
ScreenModuleEditorView "Station: ET200SP" 593x700
   GraphicView "ET200SP Stencil" at 0,50 size 593x649; Picture "ET 200SP Stencil"
   Rectangle "Interface Module Color" at 0,50 size 269x650
      Appearance <- "Interface.IM.bg"
   Rectangle "DQ 01 Module Color" at 268,50 size 95x344
      Appearance <- "Interface.DQ01.bg"
   Rectangle "DQ 01 Terminal Color" at 268,390 size 96x271
      Appearance <- "Interface.DQ01.bgTem"
   Rectangle "DQ 02 Module Color" at 363,50 size 96x344
      Appearance <- "Interface.DQ02.bg"
   Rectangle "DQ 02 Terminal Color" at 364,390 size 95x271
      Appearance <- "Interface.DQ02.bgTem"
   Rectangle "DQ 03 Module Color" at 458,50 size 95x344
      Appearance <- "Interface.DQ03.bg"
   Rectangle "DQ 03 Terminal Color" at 458,390 size 95x271
      Appearance <- "Interface.DQ03.bgTem"
   Rectangle "Server Module Color" at 552,50 size 40x343
      Appearance <- "Interface.serverModule.bg"
   Rectangle "IM Run LED" at 165,102 size 9x8
      Appearance <- "Interface.IM.run"
   Rectangle "IM Error LED" at 178,102 size 9x8
      Appearance <- "Interface.IM.error"
   Rectangle "IM Maintenance LED" at 193,102 size 9x8
      Appearance <- "Interface.IM.maint"
   Rectangle "IM Link 1 LED" at 146,295 size 9x8
      Appearance <- "Interface.IM.lnk01"
   Rectangle "IM Link 2 LED" at 146,313 size 9x8
      Appearance <- "Interface.IM.lnk02"
   Rectangle "IM Power LED" at 164,379 size 9x8
      Appearance <- "Interface.IM.pwr"
   Rectangle "DQ 01 Diag LED" at 274,102 size 9x8
      Appearance <- "Interface.DQ01.diag"
   Rectangle "DQ 01 Output LED x.0" at 274,295 size 9x8
      Appearance <- "Interface.DQ01.x0"
   Rectangle "DQ 01 Output LED x.1" at 305,295 size 9x8
      Appearance <- "Interface.DQ01.x1"
   Rectangle "DQ 01 Output LED x.2" at 274,306 size 9x8
      Appearance <- "Interface.DQ01.x2"
   Rectangle "DQ 01 Output LED x.3" at 305,306 size 9x8
      Appearance <- "Interface.DQ01.x3"
   Rectangle "DQ 01 Output LED x.4" at 274,317 size 9x8
      Appearance <- "Interface.DQ01.x4"
   Rectangle "DQ 01 Output LED x.5" at 305,317 size 9x8
      Appearance <- "Interface.DQ01.x5"
   Rectangle "DQ 01 Output LED x.6" at 274,328 size 9x8
      Appearance <- "Interface.DQ01.x6"
   Rectangle "DQ 01 Output LED x.7" at 305,328 size 9x8
      Appearance <- "Interface.DQ01.x7"
   Rectangle "DQ 01 Power LED" at 275,379 size 9x8
      Appearance <- "Interface.DQ01.pwr"
   Rectangle "DQ 02 Diag LED" at 369,102 size 9x8
      Appearance <- "Interface.DQ02.diag"
   Rectangle "DQ 02 Output LED x.0" at 369,295 size 9x8
      Appearance <- "Interface.DQ02.x0"
   Rectangle "DQ 02 Output LED x.1" at 400,295 size 9x8
      Appearance <- "Interface.DQ02.x1"
   Rectangle "DQ 02 Output LED x.2" at 369,306 size 9x8
      Appearance <- "Interface.DQ02.x2"
   Rectangle "DQ 02 Output LED x.3" at 400,306 size 9x8
      Appearance <- "Interface.DQ02.x3"
   Rectangle "DQ 02 Output LED x.4" at 369,317 size 9x8
      Appearance <- "Interface.DQ02.x4"
   Rectangle "DQ 02 Output LED x.5" at 400,317 size 9x8
      Appearance <- "Interface.DQ02.x5"
   Rectangle "DQ 02 Output LED x.6" at 369,328 size 9x8
      Appearance <- "Interface.DQ02.x6"
   Rectangle "DQ 02 Output LED x.7" at 400,328 size 9x8
      Appearance <- "Interface.DQ02.x7"
   Rectangle "DQ 02 Power LED" at 368,379 size 9x8
      Appearance <- "Interface.DQ02.pwr"
   Rectangle "DQ 03 Diag LED" at 464,102 size 9x8
      Appearance <- "Interface.DQ03.diag"
   Rectangle "DQ 03 Output LED x.0" at 464,295 size 9x8
      Appearance <- "Interface.DQ03.x0"
   Rectangle "DQ 03 Output LED x.1" at 495,295 size 9x8
      Appearance <- "Interface.DQ03.x1"
   Rectangle "DQ 03 Output LED x.2" at 464,306 size 9x8
      Appearance <- "Interface.DQ03.x2"
   Rectangle "DQ 03 Output LED x.3" at 495,306 size 9x8
      Appearance <- "Interface.DQ03.x3"
   Rectangle "DQ 03 Output LED x.4" at 464,317 size 9x8
      Appearance <- "Interface.DQ03.x4"
   Rectangle "DQ 03 Output LED x.5" at 495,317 size 9x8
      Appearance <- "Interface.DQ03.x5"
   Rectangle "DQ 03 Output LED x.6" at 464,328 size 9x8
      Appearance <- "Interface.DQ03.x6"
   Rectangle "DQ 03 Output LED x.7" at 495,328 size 9x8
      Appearance <- "Interface.DQ03.x7"
   Rectangle "DQ 03 Power LED" at 463,379 size 9x8
      Appearance <- "Interface.DQ03.pwr"
   Button "Dismiss PB" at 0,0 size 593x700; TextOff 'Text'
   TextField "PN Name" at 0,0 size 593x50; Text 'Text'
      Appearance <- "Interface.profinetName.animate"
*)

(* ===== HMI "HMI_RT_1" =====

ScreenModuleEditorView "Station: ET200SP" 603x710
   Rectangle "Interface Module Color" at 5,55 size 269x650
      Appearance <- "Interface.IM.bg"
   Rectangle "DQ 01 Module Color" at 273,55 size 95x344
      Appearance <- "Interface.DQ01.bg"
   Rectangle "DQ 01 Terminal Color" at 273,395 size 96x271
      Appearance <- "Interface.DQ01.bgTem"
   Rectangle "DQ 02 Module Color" at 368,55 size 96x344
      Appearance <- "Interface.DQ02.bg"
   Rectangle "DQ 02 Terminal Color" at 369,395 size 95x271
      Appearance <- "Interface.DQ02.bgTem"
   Rectangle "DQ 03 Module Color" at 463,55 size 95x344
      Appearance <- "Interface.DQ03.bg"
   Rectangle "DQ 03 Terminal Color" at 463,395 size 95x271
      Appearance <- "Interface.DQ03.bgTem"
   Rectangle "Server Module Color" at 557,55 size 40x343
      Appearance <- "Interface.serverModule.bg"
   Rectangle "IM Run LED" at 170,107 size 9x8
      Appearance <- "Interface.IM.run"
   Rectangle "IM Error LED" at 183,107 size 9x8
      Appearance <- "Interface.IM.error"
   Rectangle "IM Maintenance LED" at 198,107 size 9x8
      Appearance <- "Interface.IM.maint"
   Rectangle "IM Link 1 LED" at 151,300 size 9x8
      Appearance <- "Interface.IM.lnk01"
   Rectangle "IM Link 2 LED" at 151,318 size 9x8
      Appearance <- "Interface.IM.lnk02"
   Rectangle "IM Power LED" at 169,384 size 9x8
      Appearance <- "Interface.IM.pwr"
   Rectangle "DQ 01 Diag LED" at 279,107 size 9x8
      Appearance <- "Interface.DQ01.diag"
   Rectangle "DQ 01 Output LED x.0" at 279,300 size 9x8
      Appearance <- "Interface.DQ01.x0"
   Rectangle "DQ 01 Output LED x.1" at 310,300 size 9x8
      Appearance <- "Interface.DQ01.x1"
   Rectangle "DQ 01 Output LED x.2" at 279,311 size 9x8
      Appearance <- "Interface.DQ01.x2"
   Rectangle "DQ 01 Output LED x.3" at 310,311 size 9x8
      Appearance <- "Interface.DQ01.x3"
   Rectangle "DQ 01 Output LED x.4" at 279,322 size 9x8
      Appearance <- "Interface.DQ01.x4"
   Rectangle "DQ 01 Output LED x.5" at 310,322 size 9x8
      Appearance <- "Interface.DQ01.x5"
   Rectangle "DQ 01 Output LED x.6" at 279,333 size 9x8
      Appearance <- "Interface.DQ01.x6"
   Rectangle "DQ 01 Output LED x.7" at 310,333 size 9x8
      Appearance <- "Interface.DQ01.x7"
   Rectangle "DQ 01 Power LED" at 280,384 size 9x8
      Appearance <- "Interface.DQ01.pwr"
   Rectangle "DQ 02 Diag LED" at 374,107 size 9x8
      Appearance <- "Interface.DQ02.diag"
   Rectangle "DQ 02 Output LED x.0" at 374,300 size 9x8
      Appearance <- "Interface.DQ02.x0"
   Rectangle "DQ 02 Output LED x.1" at 405,300 size 9x8
      Appearance <- "Interface.DQ02.x1"
   Rectangle "DQ 02 Output LED x.2" at 374,311 size 9x8
      Appearance <- "Interface.DQ02.x2"
   Rectangle "DQ 02 Output LED x.3" at 405,311 size 9x8
      Appearance <- "Interface.DQ02.x3"
   Rectangle "DQ 02 Output LED x.4" at 374,322 size 9x8
      Appearance <- "Interface.DQ02.x4"
   Rectangle "DQ 02 Output LED x.5" at 405,322 size 9x8
      Appearance <- "Interface.DQ02.x5"
   Rectangle "DQ 02 Output LED x.6" at 374,333 size 9x8
      Appearance <- "Interface.DQ02.x6"
   Rectangle "DQ 02 Output LED x.7" at 405,333 size 9x8
      Appearance <- "Interface.DQ02.x7"
   Rectangle "DQ 02 Power LED" at 373,384 size 9x8
      Appearance <- "Interface.DQ02.pwr"
   Rectangle "DQ 03 Diag LED" at 469,107 size 9x8
      Appearance <- "Interface.DQ03.diag"
   Rectangle "DQ 03 Output LED x.0" at 469,300 size 9x8
      Appearance <- "Interface.DQ03.x0"
   Rectangle "DQ 03 Output LED x.1" at 500,300 size 9x8
      Appearance <- "Interface.DQ03.x1"
   Rectangle "DQ 03 Output LED x.2" at 469,311 size 9x8
      Appearance <- "Interface.DQ03.x2"
   Rectangle "DQ 03 Output LED x.3" at 500,311 size 9x8
      Appearance <- "Interface.DQ03.x3"
   Rectangle "DQ 03 Output LED x.4" at 469,322 size 9x8
      Appearance <- "Interface.DQ03.x4"
   Rectangle "DQ 03 Output LED x.5" at 500,322 size 9x8
      Appearance <- "Interface.DQ03.x5"
   Rectangle "DQ 03 Output LED x.6" at 469,333 size 9x8
      Appearance <- "Interface.DQ03.x6"
   Rectangle "DQ 03 Output LED x.7" at 500,333 size 9x8
      Appearance <- "Interface.DQ03.x7"
   Rectangle "DQ 03 Power LED" at 468,384 size 9x8
      Appearance <- "Interface.DQ03.pwr"
   GraphicView "ET200SP Stencil" at 5,55 size 593x649; Picture "ET 200SP Stencil"
   Button "Dismiss PB" at 5,5 size 593x700; TextOff 'Text'
   TextField "PN Name" at 5,5 size 593x50; Text 'Text'
      Appearance <- "Interface.profinetName.animate"
*)

(* ===== HMI "HMI_RT_1" =====

ScreenModuleEditorView "Station: KP8" 428x710
   GraphicView "KP8 Stencil" at 5,55 size 418x650; Picture "KP8 Rear View Stencil"
      Appearance <- "Interface.stencilBackground"
   TextField "PN Name Label" at 5,5 size 418x50; Text 'Text'
      Appearance <- "Interface.profinetName.animate"
   Rectangle "X1P1 Transmit" at 195,536 size 12x16
      Appearance <- "Interface.X1P1.transmit"
   Rectangle "X1P1 Receive" at 195,576 size 12x16
      Appearance <- "Interface.X1P1.receive"
   Rectangle "X1P2 Transmit" at 286,535 size 12x16
      Appearance <- "Interface.X1P2.transmit"
   Rectangle "X1P2 Receive" at 286,575 size 12x16
      Appearance <- "Interface.X1P2.receive"
   Rectangle "KP8 Background" at 5,55 size 418x650
      Appearance <- "Interface.profinetName.animate"
   Button "Dissmiss PB" at 5,5 size 418x700; TextOff 'Text'
*)

(* ===== HMI "HMI_RT_1" =====

ScreenModuleEditorView "Station: ET200SP" 603x710
   TextField "PN Name" at 5,5 size 593x50; Text 'Text'
      Appearance <- "Interface.profinetName.animate"
   Rectangle "Interface Module Color" at 5,55 size 269x650
      Appearance <- "Interface.IM.bg"
   Rectangle "DQ 01 Module Color" at 273,55 size 95x344
      Appearance <- "Interface.DQ01.bg"
   Rectangle "DQ 01 Terminal Color" at 273,395 size 96x271
      Appearance <- "Interface.DQ01.bgTem"
   Rectangle "DQ 02 Module Color" at 368,55 size 96x344
      Appearance <- "Interface.DQ02.bg"
   Rectangle "DQ 02 Terminal Color" at 369,395 size 95x271
      Appearance <- "Interface.DQ02.bgTem"
   Rectangle "DQ 03 Module Color" at 463,55 size 95x344
      Appearance <- "Interface.DQ03.bg"
   Rectangle "DQ 03 Terminal Color" at 463,395 size 95x271
      Appearance <- "Interface.DQ03.bgTem"
   Rectangle "Server Module Color" at 557,55 size 40x343
      Appearance <- "Interface.serverModule.bg"
   Rectangle "IM Run LED" at 170,107 size 9x8
      Appearance <- "Interface.IM.run"
   Rectangle "IM Error LED" at 183,107 size 9x8
      Appearance <- "Interface.IM.error"
   Rectangle "IM Maintenance LED" at 198,107 size 9x8
      Appearance <- "Interface.IM.maint"
   Rectangle "IM Link 1 LED" at 151,300 size 9x8
      Appearance <- "Interface.IM.lnk01"
   Rectangle "IM Link 2 LED" at 151,318 size 9x8
      Appearance <- "Interface.IM.lnk02"
   Rectangle "IM Power LED" at 169,384 size 9x8
      Appearance <- "Interface.IM.pwr"
   Rectangle "DQ 01 Diag LED" at 279,107 size 9x8
      Appearance <- "Interface.DQ01.diag"
   Rectangle "DQ 01 Output LED x.0" at 279,300 size 9x8
      Appearance <- "Interface.DQ01.x0"
   Rectangle "DQ 01 Output LED x.1" at 310,300 size 9x8
      Appearance <- "Interface.DQ01.x1"
   Rectangle "DQ 01 Output LED x.2" at 279,311 size 9x8
      Appearance <- "Interface.DQ01.x2"
   Rectangle "DQ 01 Output LED x.3" at 310,311 size 9x8
      Appearance <- "Interface.DQ01.x3"
   Rectangle "DQ 01 Output LED x.4" at 279,322 size 9x8
      Appearance <- "Interface.DQ01.x4"
   Rectangle "DQ 01 Output LED x.5" at 310,322 size 9x8
      Appearance <- "Interface.DQ01.x5"
   Rectangle "DQ 01 Output LED x.6" at 279,333 size 9x8
      Appearance <- "Interface.DQ01.x6"
   Rectangle "DQ 01 Output LED x.7" at 310,333 size 9x8
      Appearance <- "Interface.DQ01.x7"
   Rectangle "DQ 01 Power LED" at 280,384 size 9x8
      Appearance <- "Interface.DQ01.pwr"
   Rectangle "DQ 02 Diag LED" at 374,107 size 9x8
      Appearance <- "Interface.DQ02.diag"
   Rectangle "DQ 02 Output LED x.0" at 374,300 size 9x8
      Appearance <- "Interface.DQ02.x0"
   Rectangle "DQ 02 Output LED x.1" at 405,300 size 9x8
      Appearance <- "Interface.DQ02.x1"
   Rectangle "DQ 02 Output LED x.2" at 374,311 size 9x8
      Appearance <- "Interface.DQ02.x2"
   Rectangle "DQ 02 Output LED x.3" at 405,311 size 9x8
      Appearance <- "Interface.DQ02.x3"
   Rectangle "DQ 02 Output LED x.4" at 374,322 size 9x8
      Appearance <- "Interface.DQ02.x4"
   Rectangle "DQ 02 Output LED x.5" at 405,322 size 9x8
      Appearance <- "Interface.DQ02.x5"
   Rectangle "DQ 02 Output LED x.6" at 374,333 size 9x8
      Appearance <- "Interface.DQ02.x6"
   Rectangle "DQ 02 Output LED x.7" at 405,333 size 9x8
      Appearance <- "Interface.DQ02.x7"
   Rectangle "DQ 02 Power LED" at 373,384 size 9x8
      Appearance <- "Interface.DQ02.pwr"
   Rectangle "DQ 03 Diag LED" at 469,107 size 9x8
      Appearance <- "Interface.DQ03.diag"
   Rectangle "DQ 03 Output LED x.0" at 469,300 size 9x8
      Appearance <- "Interface.DQ03.x0"
   Rectangle "DQ 03 Output LED x.1" at 500,300 size 9x8
      Appearance <- "Interface.DQ03.x1"
   Rectangle "DQ 03 Output LED x.2" at 469,311 size 9x8
      Appearance <- "Interface.DQ03.x2"
   Rectangle "DQ 03 Output LED x.3" at 500,311 size 9x8
      Appearance <- "Interface.DQ03.x3"
   Rectangle "DQ 03 Output LED x.4" at 469,322 size 9x8
      Appearance <- "Interface.DQ03.x4"
   Rectangle "DQ 03 Output LED x.5" at 500,322 size 9x8
      Appearance <- "Interface.DQ03.x5"
   Rectangle "DQ 03 Output LED x.6" at 469,333 size 9x8
      Appearance <- "Interface.DQ03.x6"
   Rectangle "DQ 03 Output LED x.7" at 500,333 size 9x8
      Appearance <- "Interface.DQ03.x7"
   Rectangle "DQ 03 Power LED" at 468,384 size 9x8
      Appearance <- "Interface.DQ03.pwr"
   GraphicView "ET200SP Stencil" at 5,55 size 593x649; Picture "ET 200SP Stencil"
   Button "Dismiss PB" at 5,5 size 593x700; TextOff 'Text'
*)

(* ===== HMI "HMI_RT_3" =====
system functions are stored by id; their names below are inferred from use
connection "cv04": ETHERNET, SMART_S7_1500_OMS

HMI tags "Default tag table"
   "station" : HMI Station: Compressed = PLC "HMI Stations: HMI Data".me[3] AT %DB1.DBW0, 100 ms

Template "Current Menu Selection" 480x800
   IOField "Menu Select Label" at 6,5 size 470x154; FormatPattern ????????????????????????????????????????????????????????????
      Appearance <- "[0]"
      Visibility <- "[0]"
      ProcessValue <- "[0]"
   Button "PB Menu Select" at 6,5 size 470x154; TextOff 'Text'
      on Release: ActivateScreen("02 Menu Select", 0)
      on Press: function_b14e0dd5("pb", 0)

screen "01 Part Select" 480x800, template "Current Menu Selection"
   Button "B7" at 6,164 size 233x154; TextOff 'Text'
      on Press: function_b14e0dd5("pbs", 7)
      Visibility <- "[7]"
   Button "B6" at 6,323 size 233x154; TextOff 'Text'
      on Press: function_b14e0dd5("pbs", 6)
      Visibility <- "[6]"
   Button "B5" at 6,482 size 233x154; TextOff 'Text'
      on Press: function_b14e0dd5("pbs", 5)
      Visibility <- "[5]"
   Button "B4" at 6,641 size 233x154; TextOff 'Text'
      on Press: function_b14e0dd5("pbs", 4)
      Visibility <- "[4]"
   Button "B3" at 244,164 size 232x154; TextOff 'Text'
      on Press: function_b14e0dd5("pbs", 3)
      Visibility <- "[3]"
   Button "B2" at 244,323 size 232x154; TextOff 'Text'
      on Press: function_b14e0dd5("pbs", 2)
      Visibility <- "[2]"
   Button "B1" at 244,482 size 232x154; TextOff 'Text'
      on Press: function_b14e0dd5("pbs", 1)
      Visibility <- "[1]"
   Button "B0" at 244,641 size 232x154; TextOff 'Text'
      on Press: function_b14e0dd5("pbs", 0)
   IOField "B7 Label" at 6,164 size 233x154; FormatPattern ????????????????????????????????????????
      Appearance <- "[7]"
      ProcessValue <- "[7]"
      Visibility <- "[7]"
   IOField "B6 Label" at 6,323 size 233x154; FormatPattern ????????????????????????????????????????
      Appearance <- "[6]"
      ProcessValue <- "[6]"
      Visibility <- "[6]"
   IOField "B5 Label" at 6,482 size 233x154; FormatPattern ????????????????????????????????????????
      Appearance <- "[5]"
      ProcessValue <- "[5]"
      Visibility <- "[5]"
   IOField "B4 Label" at 6,641 size 233x154; FormatPattern ????????????????????????????????????????
      Appearance <- "[4]"
      ProcessValue <- "[4]"
      Visibility <- "[4]"
   IOField "B3 Label" at 244,164 size 232x154; FormatPattern ????????????????????????????????????????
      Appearance <- "[3]"
      ProcessValue <- "[3]"
      Visibility <- "[3]"
   IOField "B2 Label" at 244,323 size 232x154; FormatPattern ????????????????????????????????????????
      Appearance <- "[2]"
      ProcessValue <- "[2]"
      Visibility <- "[2]"
   IOField "B1 Label" at 244,482 size 232x154; FormatPattern ????????????????????????????????????????
      Appearance <- "[1]"
      ProcessValue <- "[1]"
      Visibility <- "[1]"
   IOField "B0 Label" at 244,641 size 232x154; FormatPattern ????????????????????????????????????????
      Appearance <- "[0]"
      ProcessValue <- "[0]"
      Visibility <- "[0]"

screen "02 Menu Select" 480x800, template "Current Menu Selection"
   Button "Top" at 375,164 size 100x101; TextOff 'Text'; PictureOff "basic panel top"
      on Press: function_b14e0dd5("pbs", 0)
      Appearance <- "[0]"
      Visibility <- "[0]"
   Button "Page Up" at 375,270 size 100x101; TextOff 'Text'; PictureOff "basic panel page up"
      on Press: function_b14e0dd5("pbs", 1)
      Visibility <- "[1]"
      Appearance <- "[1]"
   Button "Line Up" at 375,376 size 100x101; TextOff 'Text'; PictureOff "basic panel line up"
      on Press: function_b14e0dd5("pbs", 2)
      Appearance <- "[2]"
      Visibility <- "[2]"
   Button "Line Down" at 375,482 size 100x101; TextOff 'Text'; PictureOff "basic panel line down"
      on Press: function_b14e0dd5("pbs", 3)
      Visibility <- "[3]"
      Appearance <- "[3]"
   Button "Page Down" at 375,588 size 100x101; TextOff 'Text'; PictureOff "basic panel page down"
      on Press: function_b14e0dd5("pbs", 4)
      Appearance <- "[4]"
      Visibility <- "[4]"
   Button "Bottom" at 375,694 size 100x101; TextOff 'Text'; PictureOff "basic panel bottom"
      on Press: function_b14e0dd5("pbs", 5)
      Visibility <- "[5]"
      Appearance <- "[5]"
   Button "pbShortSelectR00" at 5,164 size 365x101; TextOff 'Text'
      on Press: function_b14e0dd5("pbs", 6)
      on Release: ActivateScreen("01 Part Select", 0)
   Button "pbShortSelectR01" at 5,270 size 365x101; TextOff 'Text'
      on Press: function_b14e0dd5("pbs", 7)
      on Release: ActivateScreen("01 Part Select", 0)
   Button "pbShortSelectR02" at 5,376 size 365x101; TextOff 'Text'
      on Press: function_b14e0dd5("pbs", 8)
      on Release: ActivateScreen("01 Part Select", 0)
   Button "pbShortSelectR03" at 5,482 size 365x101; TextOff 'Text'
      on Press: function_b14e0dd5("pbs", 9)
      on Release: ActivateScreen("01 Part Select", 0)
   Button "pbShortSelectR04" at 5,588 size 365x101; TextOff 'Text'
      on Press: function_b14e0dd5("pbs", 10)
      on Release: ActivateScreen("01 Part Select", 0)
   Button "pbShortSelectR05" at 5,694 size 365x101; TextOff 'Text'
      on Press: function_b14e0dd5("pbs", 11)
      on Release: ActivateScreen("01 Part Select", 0)
   IOField "iofShortMenuSelectR00" at 42,166 size 325x97; FormatPattern ????????????????????????????????????????????????????????????
      ProcessValue <- "[7]"
      Visibility <- "[6]"
      Appearance <- "[6]"
   IOField "iofShortMenuSelectR01" at 42,272 size 325x97; FormatPattern ????????????????????????????????????????????????????????????
      ProcessValue <- "[9]"
      Visibility <- "[7]"
      Appearance <- "[7]"
   IOField "iofShortMenuSelectR02" at 42,378 size 325x97; FormatPattern ????????????????????????????????????????????????????????????
      ProcessValue <- "[11]"
      Visibility <- "[8]"
      Appearance <- "[8]"
   IOField "iofShortMenuSelectR03" at 42,484 size 325x97; FormatPattern ????????????????????????????????????????????????????????????
      ProcessValue <- "[13]"
      Visibility <- "[9]"
      Appearance <- "[9]"
   IOField "iofShortMenuSelectR04" at 42,590 size 325x97; FormatPattern ????????????????????????????????????????????????????????????
      ProcessValue <- "[15]"
      Visibility <- "[10]"
      Appearance <- "[10]"
   IOField "iofShortMenuSelectR05" at 42,696 size 325x97; FormatPattern ????????????????????????????????????????????????????????????
      ProcessValue <- "[17]"
      Visibility <- "[11]"
      Appearance <- "[11]"
   IOField "iofLongLabelR00" at 7,166 size 35x97; FormatPattern ????????????????????????????????????????
      ProcessValue <- "[6]"
      Visibility <- "[18]"
      Appearance <- "[18]"
   IOField "iofLongLabelR01" at 7,272 size 35x97; FormatPattern ????????????????????????????????????????
      ProcessValue <- "[8]"
      Appearance <- "[19]"
      Visibility <- "[19]"
   IOField "iofLongLabelR02" at 7,378 size 35x97; FormatPattern ????????????????????????????????????????
      ProcessValue <- "[10]"
      Appearance <- "[20]"
      Visibility <- "[20]"
   IOField "iofLongLabelR03" at 7,484 size 35x97; FormatPattern ????????????????????????????????????????
      ProcessValue <- "[12]"
      Appearance <- "[21]"
      Visibility <- "[21]"
   IOField "iofLongLabelR04" at 7,590 size 35x97; FormatPattern ????????????????????????????????????????
      ProcessValue <- "[14]"
      Visibility <- "[22]"
      Appearance <- "[22]"
   IOField "iofLongtLabelR05" at 7,696 size 35x97; FormatPattern ????????????????????????????????????????
      ProcessValue <- "[16]"
      Appearance <- "[23]"
      Visibility <- "[23]"
   IOField "brdrShortR00" at 5,164 size 365x101; FormatPattern 1
      Visibility <- "[6]"
      Appearance <- "[6]"
   IOField "brdrShortR01" at 5,270 size 365x101; FormatPattern 1
      Visibility <- "[7]"
      Appearance <- "[7]"
   IOField "brdrShortR02" at 5,376 size 365x101; FormatPattern 1
      Visibility <- "[8]"
      Appearance <- "[8]"
   IOField "brdrShortR03" at 5,482 size 365x101; FormatPattern 1
      Visibility <- "[9]"
      Appearance <- "[9]"
   IOField "brdrShortR04" at 5,588 size 365x101; FormatPattern 1
      Visibility <- "[10]"
      Appearance <- "[10]"
   IOField "brdrShortR05" at 5,694 size 365x101; FormatPattern 1
      Visibility <- "[11]"
      Appearance <- "[11]"
   IOField "brdrLongR00" at 5,164 size 470x101; FormatPattern 1
      Visibility <- "[18]"
   IOField "brdrLongR01" at 5,270 size 470x101; FormatPattern 1
      Visibility <- "[19]"
   IOField "brdrLongR02" at 5,376 size 470x101; FormatPattern 1
      Visibility <- "[20]"
   IOField "brdrLongR03" at 5,482 size 470x101; FormatPattern 1
      Visibility <- "[21]"
   IOField "brdrLongR04" at 5,588 size 470x101; FormatPattern 1
      Visibility <- "[22]"
   IOField "brdrLongR05" at 5,694 size 470x101; FormatPattern 1
      Visibility <- "[23]"
   IOField "iofLongtMenuSelectR00" at 42,166 size 430x97; FormatPattern ????????????????????????????????????????????????????????????
      ProcessValue <- "[7]"
      Visibility <- "[18]"
      Appearance <- "[18]"
   IOField "iofLongtMenuSelectR01" at 42,272 size 430x97; FormatPattern ????????????????????????????????????????????????????????????
      ProcessValue <- "[9]"
      Visibility <- "[19]"
      Appearance <- "[19]"
   IOField "iofLongtMenuSelectR02" at 42,378 size 430x97; FormatPattern ????????????????????????????????????????????????????????????
      ProcessValue <- "[11]"
      Visibility <- "[20]"
      Appearance <- "[20]"
   IOField "iofLongtMenuSelectR03" at 42,484 size 430x97; FormatPattern ????????????????????????????????????????????????????????????
      ProcessValue <- "[13]"
      Visibility <- "[21]"
      Appearance <- "[21]"
   IOField "iofLongtMenuSelectR04" at 42,590 size 430x97; FormatPattern ????????????????????????????????????????????????????????????
      ProcessValue <- "[15]"
      Visibility <- "[22]"
      Appearance <- "[22]"
   IOField "iofLongtMenuSelectR05" at 42,696 size 430x97; FormatPattern ????????????????????????????????????????????????????????????
      ProcessValue <- "[17]"
      Visibility <- "[23]"
      Appearance <- "[22]"
   Button "pbLongtSelectR00" at 5,164 size 470x101; TextOff 'Text'
      on Press: function_b14e0dd5("pbs", 6)
      Visibility <- "[18]"
      on Release: ActivateScreen("01 Part Select", 0)
   Button "pbLongtSelectR01" at 5,270 size 470x101; TextOff 'Text'
      on Press: function_b14e0dd5("pbs", 7)
      Visibility <- "[19]"
      on Release: ActivateScreen("01 Part Select", 0)
   Button "pbLongtSelectR02" at 5,376 size 470x101; TextOff 'Text'
      on Press: function_b14e0dd5("pbs", 8)
      Visibility <- "[20]"
      on Release: ActivateScreen("01 Part Select", 0)
   Button "pbLongtSelectR03" at 5,482 size 470x101; TextOff 'Text'
      on Press: function_b14e0dd5("pbs", 9)
      Visibility <- "[21]"
      on Release: ActivateScreen("01 Part Select", 0)
   Button "pbLongtSelectR04" at 5,588 size 470x101; TextOff 'Text'
      on Press: function_b14e0dd5("pbs", 10)
      Visibility <- "[22]"
      on Release: ActivateScreen("01 Part Select", 0)
   Button "pbLongtSelectR05" at 5,694 size 470x101; TextOff 'Text'
      on Press: function_b14e0dd5("pbs", 11)
      Visibility <- "[23]"
      on Release: ActivateScreen("01 Part Select", 0)
   IOField "iofShortLabelR00" at 7,166 size 35x97; FormatPattern ????????????????????????????????????????
      ProcessValue <- "[6]"
      Appearance <- "[6]"
      Visibility <- "[6]"
   IOField "iofShortLabelR01" at 7,272 size 35x97; FormatPattern ????????????????????????????????????????
      ProcessValue <- "[8]"
      Appearance <- "[7]"
      Visibility <- "[7]"
   IOField "iofShortLabelR02" at 7,378 size 35x97; FormatPattern ????????????????????????????????????????
      ProcessValue <- "[10]"
      Appearance <- "[8]"
      Visibility <- "[8]"
   IOField "iofShortLabelR03" at 7,484 size 35x97; FormatPattern ????????????????????????????????????????
      ProcessValue <- "[12]"
      Appearance <- "[9]"
      Visibility <- "[9]"
   IOField "iofShortLabelR04" at 7,590 size 35x97; FormatPattern ????????????????????????????????????????
      ProcessValue <- "[14]"
      Appearance <- "[10]"
      Visibility <- "[10]"
   IOField "iofShorttLabelR05" at 7,696 size 35x97; FormatPattern ????????????????????????????????????????
      ProcessValue <- "[16]"
      Appearance <- "[11]"
      Visibility <- "[11]"
*)

(* ===== HMI "HMI_RT_4" =====
system functions are stored by id; their names below are inferred from use
connection "cv03": ETHERNET, SMART_S7_1500_OMS

HMI tags "Default tag table"
   "station" : HMI Station: Compressed = PLC "HMI Stations: HMI Data".me[2] AT %DB1.DBW0, 100 ms

screen "01 Part Select" 480x800, template "Current Menu Selection"
   Button "B7" at 6,164 size 233x154; TextOff 'Text'
      on Press: function_b14e0dd5("pbs", 7)
      Visibility <- "[7]"
   Button "B6" at 6,323 size 233x154; TextOff 'Text'
      on Press: function_b14e0dd5("pbs", 6)
      Visibility <- "[6]"
   Button "B5" at 6,482 size 233x154; TextOff 'Text'
      on Press: function_b14e0dd5("pbs", 5)
      Visibility <- "[5]"
   Button "B4" at 6,641 size 233x154; TextOff 'Text'
      on Press: function_b14e0dd5("pbs", 4)
      Visibility <- "[4]"
   Button "B3" at 244,164 size 232x154; TextOff 'Text'
      on Press: function_b14e0dd5("pbs", 3)
      Visibility <- "[3]"
   Button "B2" at 244,323 size 232x154; TextOff 'Text'
      on Press: function_b14e0dd5("pbs", 2)
      Visibility <- "[2]"
   Button "B1" at 244,482 size 232x154; TextOff 'Text'
      on Press: function_b14e0dd5("pbs", 1)
      Visibility <- "[1]"
   Button "B0" at 244,641 size 232x154; TextOff 'Text'
      on Press: function_b14e0dd5("pbs", 0)
   IOField "B7 Label" at 6,164 size 233x154; FormatPattern ????????????????????????????????????????
      Appearance <- "[7]"
      ProcessValue <- "[7]"
      Visibility <- "[7]"
   IOField "B6 Label" at 6,323 size 233x154; FormatPattern ????????????????????????????????????????
      Appearance <- "[6]"
      ProcessValue <- "[6]"
      Visibility <- "[6]"
   IOField "B5 Label" at 6,482 size 233x154; FormatPattern ????????????????????????????????????????
      Appearance <- "[5]"
      ProcessValue <- "[5]"
      Visibility <- "[5]"
   IOField "B4 Label" at 6,641 size 233x154; FormatPattern ????????????????????????????????????????
      Appearance <- "[4]"
      ProcessValue <- "[4]"
      Visibility <- "[4]"
   IOField "B3 Label" at 244,164 size 232x154; FormatPattern ????????????????????????????????????????
      Appearance <- "[3]"
      ProcessValue <- "[3]"
      Visibility <- "[3]"
   IOField "B2 Label" at 244,323 size 232x154; FormatPattern ????????????????????????????????????????
      Appearance <- "[2]"
      ProcessValue <- "[2]"
      Visibility <- "[2]"
   IOField "B1 Label" at 244,482 size 232x154; FormatPattern ????????????????????????????????????????
      Appearance <- "[1]"
      ProcessValue <- "[1]"
      Visibility <- "[1]"
   IOField "B0 Label" at 244,641 size 232x154; FormatPattern ????????????????????????????????????????
      Appearance <- "[0]"
      ProcessValue <- "[0]"
      Visibility <- "[0]"

screen "02 Menu Select" 480x800, template "Current Menu Selection"
   Button "Top" at 375,164 size 100x101; TextOff 'Text'; PictureOff "basic panel top"
      on Press: function_b14e0dd5("pbs", 0)
      Appearance <- "[0]"
      Visibility <- "[0]"
   Button "Page Up" at 375,270 size 100x101; TextOff 'Text'; PictureOff "basic panel page up"
      on Press: function_b14e0dd5("pbs", 1)
      Visibility <- "[1]"
      Appearance <- "[1]"
   Button "Line Up" at 375,376 size 100x101; TextOff 'Text'; PictureOff "basic panel line up"
      on Press: function_b14e0dd5("pbs", 2)
      Appearance <- "[2]"
      Visibility <- "[2]"
   Button "Line Down" at 375,482 size 100x101; TextOff 'Text'; PictureOff "basic panel line down"
      on Press: function_b14e0dd5("pbs", 3)
      Visibility <- "[3]"
      Appearance <- "[3]"
   Button "Page Down" at 375,588 size 100x101; TextOff 'Text'; PictureOff "basic panel page down"
      on Press: function_b14e0dd5("pbs", 4)
      Appearance <- "[4]"
      Visibility <- "[4]"
   Button "Bottom" at 375,694 size 100x101; TextOff 'Text'; PictureOff "basic panel bottom"
      on Press: function_b14e0dd5("pbs", 5)
      Visibility <- "[5]"
      Appearance <- "[5]"
   IOField "brdrShortR00" at 5,164 size 365x101; FormatPattern 1
      Visibility <- "[6]"
      Appearance <- "[6]"
   IOField "brdrShortR01" at 5,270 size 365x101; FormatPattern 1
      Visibility <- "[7]"
      Appearance <- "[7]"
   IOField "brdrShortR02" at 5,376 size 365x101; FormatPattern 1
      Visibility <- "[8]"
      Appearance <- "[8]"
   IOField "brdrShortR03" at 5,482 size 365x101; FormatPattern 1
      Visibility <- "[9]"
      Appearance <- "[9]"
   IOField "brdrShortR04" at 5,588 size 365x101; FormatPattern 1
      Visibility <- "[10]"
      Appearance <- "[10]"
   IOField "brdrShortR05" at 5,694 size 365x101; FormatPattern 1
      Visibility <- "[11]"
      Appearance <- "[11]"
   Button "pbShortSelectR00" at 5,164 size 365x101; TextOff 'Text'
      on Release: ActivateScreen("01 Part Select", 0)
      on Press: function_b14e0dd5("pbs", 6)
   Button "pbShortSelectR01" at 5,270 size 365x101; TextOff 'Text'
      on Release: ActivateScreen("01 Part Select", 0)
      on Press: function_b14e0dd5("pbs", 7)
   Button "pbShortSelectR02" at 5,376 size 365x101; TextOff 'Text'
      on Release: ActivateScreen("01 Part Select", 0)
      on Press: function_b14e0dd5("pbs", 8)
   Button "pbShortSelectR03" at 5,482 size 365x101; TextOff 'Text'
      on Release: ActivateScreen("01 Part Select", 0)
      on Press: function_b14e0dd5("pbs", 9)
   Button "pbShortSelectR04" at 5,588 size 365x101; TextOff 'Text'
      on Release: ActivateScreen("01 Part Select", 0)
      on Press: function_b14e0dd5("pbs", 10)
   Button "pbShortSelectR05" at 5,694 size 365x101; TextOff 'Text'
      on Release: ActivateScreen("01 Part Select", 0)
      on Press: function_b14e0dd5("pbs", 11)
   IOField "brdrLongR00" at 5,164 size 470x101; FormatPattern 1
      Visibility <- "[18]"
   IOField "brdrLongR01" at 5,270 size 470x101; FormatPattern 1
      Visibility <- "[19]"
   IOField "brdrLongR02" at 5,376 size 470x101; FormatPattern 1
      Visibility <- "[20]"
   IOField "brdrLongR03" at 5,482 size 470x101; FormatPattern 1
      Visibility <- "[21]"
   IOField "brdrLongR04" at 5,588 size 470x101; FormatPattern 1
      Visibility <- "[22]"
   IOField "brdrLongR05" at 5,694 size 470x101; FormatPattern 1
      Visibility <- "[23]"
   Button "pbLongtSelectR00" at 5,164 size 470x101; TextOff 'Text'
      on Release: ActivateScreen("01 Part Select", 0)
      on Press: function_b14e0dd5("pbs", 6)
      Visibility <- "[18]"
   Button "pbLongtSelectR01" at 5,270 size 470x101; TextOff 'Text'
      on Release: ActivateScreen("01 Part Select", 0)
      on Press: function_b14e0dd5("pbs", 7)
      Visibility <- "[19]"
   Button "pbLongtSelectR02" at 5,376 size 470x101; TextOff 'Text'
      on Release: ActivateScreen("01 Part Select", 0)
      on Press: function_b14e0dd5("pbs", 8)
      Visibility <- "[20]"
   Button "pbLongtSelectR03" at 5,482 size 470x101; TextOff 'Text'
      on Release: ActivateScreen("01 Part Select", 0)
      on Press: function_b14e0dd5("pbs", 9)
      Visibility <- "[21]"
   Button "pbLongtSelectR04" at 5,588 size 470x101; TextOff 'Text'
      on Release: ActivateScreen("01 Part Select", 0)
      on Press: function_b14e0dd5("pbs", 10)
      Visibility <- "[22]"
   Button "pbLongtSelectR05" at 5,694 size 470x101; TextOff 'Text'
      on Release: ActivateScreen("01 Part Select", 0)
      on Press: function_b14e0dd5("pbs", 11)
      Visibility <- "[23]"
   IOField "iofLongtMenuSelectR00" at 42,166 size 430x97; FormatPattern ????????????????????????????????????????????????????????????
      Visibility <- "[18]"
      ProcessValue <- "[7]"
      Appearance <- "[18]"
   IOField "iofLongtMenuSelectR01" at 42,272 size 430x97; FormatPattern ????????????????????????????????????????????????????????????
      Visibility <- "[19]"
      ProcessValue <- "[9]"
      Appearance <- "[19]"
   IOField "iofLongtMenuSelectR02" at 42,378 size 430x97; FormatPattern ????????????????????????????????????????????????????????????
      Visibility <- "[20]"
      ProcessValue <- "[11]"
      Appearance <- "[20]"
   IOField "iofLongtMenuSelectR03" at 42,484 size 430x97; FormatPattern ????????????????????????????????????????????????????????????
      Visibility <- "[21]"
      ProcessValue <- "[13]"
      Appearance <- "[21]"
   IOField "iofLongtMenuSelectR04" at 42,590 size 430x97; FormatPattern ????????????????????????????????????????????????????????????
      Visibility <- "[22]"
      ProcessValue <- "[15]"
      Appearance <- "[22]"
   IOField "iofLongtMenuSelectR05" at 42,696 size 430x97; FormatPattern ????????????????????????????????????????????????????????????
      Visibility <- "[23]"
      ProcessValue <- "[17]"
      Appearance <- "[22]"
   IOField "iofLongLabelR00" at 7,166 size 35x97; FormatPattern ????????????????????????????????????????
      Visibility <- "[18]"
      ProcessValue <- "[6]"
      Appearance <- "[18]"
   IOField "iofLongLabelR01" at 7,272 size 35x97; FormatPattern ????????????????????????????????????????
      Appearance <- "[19]"
      ProcessValue <- "[8]"
      Visibility <- "[19]"
   IOField "iofLongLabelR02" at 7,378 size 35x97; FormatPattern ????????????????????????????????????????
      Appearance <- "[20]"
      ProcessValue <- "[10]"
      Visibility <- "[20]"
   IOField "iofLongLabelR03" at 7,484 size 35x97; FormatPattern ????????????????????????????????????????
      Appearance <- "[21]"
      ProcessValue <- "[12]"
      Visibility <- "[21]"
   IOField "iofLongLabelR04" at 7,590 size 35x97; FormatPattern ????????????????????????????????????????
      Visibility <- "[22]"
      ProcessValue <- "[14]"
      Appearance <- "[22]"
   IOField "iofLongtLabelR05" at 7,696 size 35x97; FormatPattern ????????????????????????????????????????
      Appearance <- "[23]"
      ProcessValue <- "[16]"
      Visibility <- "[23]"
   IOField "iofShortMenuSelectR00" at 42,166 size 325x97; FormatPattern ????????????????????????????????????????????????????????????
      Visibility <- "[6]"
      ProcessValue <- "[7]"
      Appearance <- "[6]"
   IOField "iofShortMenuSelectR01" at 42,272 size 325x97; FormatPattern ????????????????????????????????????????????????????????????
      Visibility <- "[7]"
      ProcessValue <- "[9]"
      Appearance <- "[7]"
   IOField "iofShortMenuSelectR02" at 42,378 size 325x97; FormatPattern ????????????????????????????????????????????????????????????
      Visibility <- "[8]"
      ProcessValue <- "[11]"
      Appearance <- "[8]"
   IOField "iofShortMenuSelectR03" at 42,484 size 325x97; FormatPattern ????????????????????????????????????????????????????????????
      Visibility <- "[9]"
      ProcessValue <- "[13]"
      Appearance <- "[9]"
   IOField "iofShortMenuSelectR04" at 42,590 size 325x97; FormatPattern ????????????????????????????????????????????????????????????
      Visibility <- "[10]"
      ProcessValue <- "[15]"
      Appearance <- "[10]"
   IOField "iofShortMenuSelectR05" at 42,696 size 325x97; FormatPattern ????????????????????????????????????????????????????????????
      Visibility <- "[11]"
      ProcessValue <- "[17]"
      Appearance <- "[11]"
   IOField "iofShortLabelR00" at 7,166 size 35x97; FormatPattern ????????????????????????????????????????
      Appearance <- "[6]"
      ProcessValue <- "[6]"
      Visibility <- "[6]"
   IOField "iofShortLabelR01" at 7,272 size 35x97; FormatPattern ????????????????????????????????????????
      Appearance <- "[7]"
      ProcessValue <- "[8]"
      Visibility <- "[7]"
   IOField "iofShortLabelR02" at 7,378 size 35x97; FormatPattern ????????????????????????????????????????
      Appearance <- "[8]"
      ProcessValue <- "[10]"
      Visibility <- "[8]"
   IOField "iofShortLabelR03" at 7,484 size 35x97; FormatPattern ????????????????????????????????????????
      Appearance <- "[9]"
      ProcessValue <- "[12]"
      Visibility <- "[9]"
   IOField "iofShortLabelR04" at 7,590 size 35x97; FormatPattern ????????????????????????????????????????
      Appearance <- "[10]"
      ProcessValue <- "[14]"
      Visibility <- "[10]"
   IOField "iofShorttLabelR05" at 7,696 size 35x97; FormatPattern ????????????????????????????????????????
      Appearance <- "[11]"
      ProcessValue <- "[16]"
      Visibility <- "[11]"

Template "Current Menu Selection" 480x800
   IOField "Menu Select Label" at 6,5 size 470x154; FormatPattern ????????????????????????????????????????????????????????????
      Appearance <- "[0]"
      Visibility <- "[0]"
      ProcessValue <- "[0]"
   Button "PB Menu Select" at 6,5 size 470x154; TextOff 'Text'
      on Release: ActivateScreen("02 Menu Select", 0)
      on Press: function_b14e0dd5("pb", 0)
*)

(* ===== HMI "HMI_RT_5" =====
system functions are stored by id; their names below are inferred from use
connection "cv02": ETHERNET, SMART_S7_1500_OMS

HMI tags "Default tag table"
   "station" : HMI Station: Compressed = PLC "HMI Stations: HMI Data".me[1] AT %DB1.DBW0, 100 ms

screen "01 Part Select" 480x800, template "Current Menu Selection"
   Button "B7" at 6,164 size 233x154; TextOff 'Text'
      on Press: function_b14e0dd5("pbs", 7)
      Visibility <- "[7]"
   Button "B6" at 6,323 size 233x154; TextOff 'Text'
      on Press: function_b14e0dd5("pbs", 6)
      Visibility <- "[6]"
   Button "B5" at 6,482 size 233x154; TextOff 'Text'
      on Press: function_b14e0dd5("pbs", 5)
      Visibility <- "[5]"
   Button "B4" at 6,641 size 233x154; TextOff 'Text'
      on Press: function_b14e0dd5("pbs", 4)
      Visibility <- "[4]"
   Button "B3" at 244,164 size 232x154; TextOff 'Text'
      on Press: function_b14e0dd5("pbs", 3)
      Visibility <- "[3]"
   Button "B2" at 244,323 size 232x154; TextOff 'Text'
      on Press: function_b14e0dd5("pbs", 2)
      Visibility <- "[2]"
   Button "B1" at 244,482 size 232x154; TextOff 'Text'
      on Press: function_b14e0dd5("pbs", 1)
      Visibility <- "[1]"
   Button "B0" at 244,641 size 232x154; TextOff 'Text'
      on Press: function_b14e0dd5("pbs", 0)
   IOField "B7 Label" at 6,164 size 233x154; FormatPattern ????????????????????????????????????????
      Appearance <- "[7]"
      ProcessValue <- "[7]"
      Visibility <- "[7]"
   IOField "B6 Label" at 6,323 size 233x154; FormatPattern ????????????????????????????????????????
      Appearance <- "[6]"
      ProcessValue <- "[6]"
      Visibility <- "[6]"
   IOField "B5 Label" at 6,482 size 233x154; FormatPattern ????????????????????????????????????????
      Appearance <- "[5]"
      ProcessValue <- "[5]"
      Visibility <- "[5]"
   IOField "B4 Label" at 6,641 size 233x154; FormatPattern ????????????????????????????????????????
      Appearance <- "[4]"
      ProcessValue <- "[4]"
      Visibility <- "[4]"
   IOField "B3 Label" at 244,164 size 232x154; FormatPattern ????????????????????????????????????????
      Appearance <- "[3]"
      ProcessValue <- "[3]"
      Visibility <- "[3]"
   IOField "B2 Label" at 244,323 size 232x154; FormatPattern ????????????????????????????????????????
      Appearance <- "[2]"
      ProcessValue <- "[2]"
      Visibility <- "[2]"
   IOField "B1 Label" at 244,482 size 232x154; FormatPattern ????????????????????????????????????????
      Appearance <- "[1]"
      ProcessValue <- "[1]"
      Visibility <- "[1]"
   IOField "B0 Label" at 244,641 size 232x154; FormatPattern ????????????????????????????????????????
      Appearance <- "[0]"
      ProcessValue <- "[0]"
      Visibility <- "[0]"

screen "02 Menu Select" 480x800, template "Current Menu Selection"
   Button "Top" at 375,164 size 100x101; TextOff 'Text'; PictureOff "basic panel top"
      on Press: function_b14e0dd5("pbs", 0)
      Appearance <- "[0]"
      Visibility <- "[0]"
   Button "Page Up" at 375,270 size 100x101; TextOff 'Text'; PictureOff "basic panel page up"
      on Press: function_b14e0dd5("pbs", 1)
      Visibility <- "[1]"
      Appearance <- "[1]"
   Button "Line Up" at 375,376 size 100x101; TextOff 'Text'; PictureOff "basic panel line up"
      on Press: function_b14e0dd5("pbs", 2)
      Appearance <- "[2]"
      Visibility <- "[2]"
   Button "Line Down" at 375,482 size 100x101; TextOff 'Text'; PictureOff "basic panel line down"
      on Press: function_b14e0dd5("pbs", 3)
      Visibility <- "[3]"
      Appearance <- "[3]"
   Button "Page Down" at 375,588 size 100x101; TextOff 'Text'; PictureOff "basic panel page down"
      on Press: function_b14e0dd5("pbs", 4)
      Appearance <- "[4]"
      Visibility <- "[4]"
   Button "Bottom" at 375,694 size 100x101; TextOff 'Text'; PictureOff "basic panel bottom"
      on Press: function_b14e0dd5("pbs", 5)
      Visibility <- "[5]"
      Appearance <- "[5]"
   IOField "brdrShortR00" at 5,164 size 365x101; FormatPattern 1
      Visibility <- "[6]"
      Appearance <- "[6]"
   IOField "brdrShortR01" at 5,270 size 365x101; FormatPattern 1
      Visibility <- "[7]"
      Appearance <- "[7]"
   IOField "brdrShortR02" at 5,376 size 365x101; FormatPattern 1
      Visibility <- "[8]"
      Appearance <- "[8]"
   IOField "brdrShortR03" at 5,482 size 365x101; FormatPattern 1
      Visibility <- "[9]"
      Appearance <- "[9]"
   IOField "brdrShortR04" at 5,588 size 365x101; FormatPattern 1
      Visibility <- "[10]"
      Appearance <- "[10]"
   IOField "brdrShortR05" at 5,694 size 365x101; FormatPattern 1
      Visibility <- "[11]"
      Appearance <- "[11]"
   Button "pbShortSelectR00" at 5,164 size 365x101; TextOff 'Text'
      on Release: ActivateScreen("01 Part Select", 0)
      on Press: function_b14e0dd5("pbs", 6)
   Button "pbShortSelectR01" at 5,270 size 365x101; TextOff 'Text'
      on Release: ActivateScreen("01 Part Select", 0)
      on Press: function_b14e0dd5("pbs", 7)
   Button "pbShortSelectR02" at 5,376 size 365x101; TextOff 'Text'
      on Release: ActivateScreen("01 Part Select", 0)
      on Press: function_b14e0dd5("pbs", 8)
   Button "pbShortSelectR03" at 5,482 size 365x101; TextOff 'Text'
      on Release: ActivateScreen("01 Part Select", 0)
      on Press: function_b14e0dd5("pbs", 9)
   Button "pbShortSelectR04" at 5,588 size 365x101; TextOff 'Text'
      on Release: ActivateScreen("01 Part Select", 0)
      on Press: function_b14e0dd5("pbs", 10)
   Button "pbShortSelectR05" at 5,694 size 365x101; TextOff 'Text'
      on Release: ActivateScreen("01 Part Select", 0)
      on Press: function_b14e0dd5("pbs", 11)
   IOField "brdrLongR00" at 5,164 size 470x101; FormatPattern 1
      Visibility <- "[18]"
   IOField "brdrLongR01" at 5,270 size 470x101; FormatPattern 1
      Visibility <- "[19]"
   IOField "brdrLongR02" at 5,376 size 470x101; FormatPattern 1
      Visibility <- "[20]"
   IOField "brdrLongR03" at 5,482 size 470x101; FormatPattern 1
      Visibility <- "[21]"
   IOField "brdrLongR04" at 5,588 size 470x101; FormatPattern 1
      Visibility <- "[22]"
   IOField "brdrLongR05" at 5,694 size 470x101; FormatPattern 1
      Visibility <- "[23]"
   Button "pbLongtSelectR00" at 5,164 size 470x101; TextOff 'Text'
      on Release: ActivateScreen("01 Part Select", 0)
      on Press: function_b14e0dd5("pbs", 6)
      Visibility <- "[18]"
   Button "pbLongtSelectR01" at 5,270 size 470x101; TextOff 'Text'
      on Release: ActivateScreen("01 Part Select", 0)
      on Press: function_b14e0dd5("pbs", 7)
      Visibility <- "[19]"
   Button "pbLongtSelectR02" at 5,376 size 470x101; TextOff 'Text'
      on Release: ActivateScreen("01 Part Select", 0)
      on Press: function_b14e0dd5("pbs", 8)
      Visibility <- "[20]"
   Button "pbLongtSelectR03" at 5,482 size 470x101; TextOff 'Text'
      on Release: ActivateScreen("01 Part Select", 0)
      on Press: function_b14e0dd5("pbs", 9)
      Visibility <- "[21]"
   Button "pbLongtSelectR04" at 5,588 size 470x101; TextOff 'Text'
      on Release: ActivateScreen("01 Part Select", 0)
      on Press: function_b14e0dd5("pbs", 10)
      Visibility <- "[22]"
   Button "pbLongtSelectR05" at 5,694 size 470x101; TextOff 'Text'
      on Release: ActivateScreen("01 Part Select", 0)
      on Press: function_b14e0dd5("pbs", 11)
      Visibility <- "[23]"
   IOField "iofLongtMenuSelectR00" at 42,166 size 430x97; FormatPattern ????????????????????????????????????????????????????????????
      Visibility <- "[18]"
      ProcessValue <- "[7]"
      Appearance <- "[18]"
   IOField "iofLongtMenuSelectR01" at 42,272 size 430x97; FormatPattern ????????????????????????????????????????????????????????????
      Visibility <- "[19]"
      ProcessValue <- "[9]"
      Appearance <- "[19]"
   IOField "iofLongtMenuSelectR02" at 42,378 size 430x97; FormatPattern ????????????????????????????????????????????????????????????
      Visibility <- "[20]"
      ProcessValue <- "[11]"
      Appearance <- "[20]"
   IOField "iofLongtMenuSelectR03" at 42,484 size 430x97; FormatPattern ????????????????????????????????????????????????????????????
      Visibility <- "[21]"
      ProcessValue <- "[13]"
      Appearance <- "[21]"
   IOField "iofLongtMenuSelectR04" at 42,590 size 430x97; FormatPattern ????????????????????????????????????????????????????????????
      Visibility <- "[22]"
      ProcessValue <- "[15]"
      Appearance <- "[22]"
   IOField "iofLongtMenuSelectR05" at 42,696 size 430x97; FormatPattern ????????????????????????????????????????????????????????????
      Visibility <- "[23]"
      ProcessValue <- "[17]"
      Appearance <- "[22]"
   IOField "iofLongLabelR00" at 7,166 size 35x97; FormatPattern ????????????????????????????????????????
      Visibility <- "[18]"
      ProcessValue <- "[6]"
      Appearance <- "[18]"
   IOField "iofLongLabelR01" at 7,272 size 35x97; FormatPattern ????????????????????????????????????????
      Appearance <- "[19]"
      ProcessValue <- "[8]"
      Visibility <- "[19]"
   IOField "iofLongLabelR02" at 7,378 size 35x97; FormatPattern ????????????????????????????????????????
      Appearance <- "[20]"
      ProcessValue <- "[10]"
      Visibility <- "[20]"
   IOField "iofLongLabelR03" at 7,484 size 35x97; FormatPattern ????????????????????????????????????????
      Appearance <- "[21]"
      ProcessValue <- "[12]"
      Visibility <- "[21]"
   IOField "iofLongLabelR04" at 7,590 size 35x97; FormatPattern ????????????????????????????????????????
      Visibility <- "[22]"
      ProcessValue <- "[14]"
      Appearance <- "[22]"
   IOField "iofLongtLabelR05" at 7,696 size 35x97; FormatPattern ????????????????????????????????????????
      Appearance <- "[23]"
      ProcessValue <- "[16]"
      Visibility <- "[23]"
   IOField "iofShortMenuSelectR00" at 42,166 size 325x97; FormatPattern ????????????????????????????????????????????????????????????
      Visibility <- "[6]"
      ProcessValue <- "[7]"
      Appearance <- "[6]"
   IOField "iofShortMenuSelectR01" at 42,272 size 325x97; FormatPattern ????????????????????????????????????????????????????????????
      Visibility <- "[7]"
      ProcessValue <- "[9]"
      Appearance <- "[7]"
   IOField "iofShortMenuSelectR02" at 42,378 size 325x97; FormatPattern ????????????????????????????????????????????????????????????
      Visibility <- "[8]"
      ProcessValue <- "[11]"
      Appearance <- "[8]"
   IOField "iofShortMenuSelectR03" at 42,484 size 325x97; FormatPattern ????????????????????????????????????????????????????????????
      Visibility <- "[9]"
      ProcessValue <- "[13]"
      Appearance <- "[9]"
   IOField "iofShortMenuSelectR04" at 42,590 size 325x97; FormatPattern ????????????????????????????????????????????????????????????
      Visibility <- "[10]"
      ProcessValue <- "[15]"
      Appearance <- "[10]"
   IOField "iofShortMenuSelectR05" at 42,696 size 325x97; FormatPattern ????????????????????????????????????????????????????????????
      Visibility <- "[11]"
      ProcessValue <- "[17]"
      Appearance <- "[11]"
   IOField "iofShortLabelR00" at 7,166 size 35x97; FormatPattern ????????????????????????????????????????
      Appearance <- "[6]"
      ProcessValue <- "[6]"
      Visibility <- "[6]"
   IOField "iofShortLabelR01" at 7,272 size 35x97; FormatPattern ????????????????????????????????????????
      Appearance <- "[7]"
      ProcessValue <- "[8]"
      Visibility <- "[7]"
   IOField "iofShortLabelR02" at 7,378 size 35x97; FormatPattern ????????????????????????????????????????
      Appearance <- "[8]"
      ProcessValue <- "[10]"
      Visibility <- "[8]"
   IOField "iofShortLabelR03" at 7,484 size 35x97; FormatPattern ????????????????????????????????????????
      Appearance <- "[9]"
      ProcessValue <- "[12]"
      Visibility <- "[9]"
   IOField "iofShortLabelR04" at 7,590 size 35x97; FormatPattern ????????????????????????????????????????
      Appearance <- "[10]"
      ProcessValue <- "[14]"
      Visibility <- "[10]"
   IOField "iofShorttLabelR05" at 7,696 size 35x97; FormatPattern ????????????????????????????????????????
      Appearance <- "[11]"
      ProcessValue <- "[16]"
      Visibility <- "[11]"

Template "Current Menu Selection" 480x800
   IOField "Menu Select Label" at 6,5 size 470x154; FormatPattern ????????????????????????????????????????????????????????????
      Appearance <- "[0]"
      Visibility <- "[0]"
      ProcessValue <- "[0]"
   Button "PB Menu Select" at 6,5 size 470x154; TextOff 'Text'
      on Release: ActivateScreen("02 Menu Select", 0)
      on Press: function_b14e0dd5("pb", 0)
*)

(* ===== HMI "HMI_RT_6" =====
system functions are stored by id; their names below are inferred from use
connection "cv01": ETHERNET, SMART_S7_1500_OMS

